// TIA Portal project "g" (V14)

(* hardware
DEVICE "S7-1200 station_1"  S7-1200 Station
   slot 0: "Rack_0"  S7-1200 Rack  Rack  V1.0
   slot 1: "PLC_1_test_mb_og_utv"  CPU 1217C DC/DC/DC  6ES7 217-1AG40-0XB0  V4.2
   slot 2: "DI 16x24VDC_1"  6ES7 221-1BH32-0XB0  V2.0
   slot 3: "CB 1241 (RS485)"  CB 1241 (RS485)  6ES7 241-1CH30-1XB0  V1.0
DEVICE "S7-1200 station_6"  S7-1200 Station
   slot 0: "Rack_0"  S7-1200 Rack  Rack  V1.0
   slot 1: "slib"  CPU 1211C DC/DC/DC  6ES7 211-1AE40-0XB0  V4.2
   slot 3: "CB 1241 (RS485)"  CB 1241 (RS485)  6ES7 241-1CH30-1XB0  V1.0
DEVICE "HMI"  TP900 Comfort
   slot 0: "TP900 Comfort"  TP900 Comfort  6AV2 124-0JC01-0AX0  14.0.1.0
   slot 1: "HMI_RT_2"  TP900 Comfort  6AV2 124-0JC01-0AX0  14.0.1.0
   slot 5: "HMI_2.IE_CP_1"  PROFINET Interface  14.0.1.0
      slot 1: "PROFINET Interface_1"  PROFINET Interface
         slot 1: "Port_1"  Port
         slot 2: "Port_2"  Port
   slot 7: "HMI_2.MPI/DP_CP_1"  MPI/DP Interface  14.0.1.0
DEVICE "S7-1200 station_2"  S7-1200 Station
   slot 0: "Rack_0"  S7-1200 Rack  Rack  V1.0
   slot 1: "PLC_1"  CPU 1211C DC/DC/DC  6ES7 211-1AE40-0XB0  V4.2
   slot 3: "CB 1241 (RS485)"  CB 1241 (RS485)  6ES7 241-1CH30-1XB0  V1.0
*)

// ===== PLC "PLC_1_test_mb_og_utv"  CPU 1217C DC/DC/DC =====

VAR_GLOBAL   // PLC tag table "Default tag table"
   "my_special_tag_name" AT %IW0 : Int;
   "tt" AT %I0.0 : Bool;
END_VAR

TYPE "mb_station_block_udt"
   STRUCT
      conf : Struct   // Configuration
         disable : Bool;   // Skip all queries
         read_only : Bool;   // Skip all write queries. (fc 5,6,15,16)
         max_comm_error : USInt := 2;   // Repeating erros before communication_error flag is set
         exec_x_quries : USInt := 1;   // Number of queries to be exec. at each loop.
      END_STRUCT;
      out : Struct   // Outputs
         error : Bool;   // All errors, including communication errors
         error_comm : Bool;   // only communication errors
         finnish : Bool;   // qid is handed over to next device.
      END_STRUCT;
      log : Struct   // Logging for development and debugging.
         connected_time : DTL;   // The time the device was connected to the bus
         disconnected_time : DTL;   // The time, if a device was disconnected to the bus
         done_cnt : UDInt;   // Successfully queries counter for this device
         error_comm_cnt : UDInt;   // Communication erros cnt.
         error_exception_cnt : UDInt;   // Failed queries counter for this device
         error_status : Word;   // Status code from mb_master or mb_client
         error_data_addr : UDInt;   // d_addr for last failed querie; handy for troubleshooting
      END_STRUCT;
      z : Struct   // Internal states.
         header_qid : UInt;   // qid value at device header
         comm_err_cnt : USInt;   // Repeating communication errors
         exec_cnt : USInt;   // Numb. of exec. q. this loop
         offset_qid : UInt := 1;   // Device query id.
         err_hold : Bool;   // Help var for .out.error
      END_STRUCT;
   END_STRUCT;
END_TYPE

// folder: mb_test

DATA_BLOCK "test_mb_t1_DB"   // DB1
{ S7_Optimized_Access := 'TRUE' }
VERSION : 0.1
// stored: InstanceOfName test_mb_1
"test_mb_1"
BEGIN
END_DATA_BLOCK

// folder: (top level)

FUNCTION_BLOCK "_read little"   // FB1, SCL
{ S7_Optimized_Access := 'TRUE' }
VERSION : 0.1
   VAR_INPUT
      mb_addr : USInt;
   END_VAR
   VAR_IN_OUT
      mb_query : "mb_query";
   END_VAR
   VAR
      sb : "mb_station_block_udt";
      data1 : Real;
      data2 : Real;
      data3 : Real;
      dommy : Bool;
      err : Int;
      pos : DInt;
   END_VAR
BEGIN

   #mb_query(mb_addr := 123,
             mode := #mb_query.c.read.holding_reg,
             data_addr := 12345,
             data_ptr := #dommy);

   IF #mb_query.Done THEN

       // #pos := "mb_pos"(mb_query := #mb_query, addr := 12345);
       #pos := UDINT_TO_DINT(12354 - #mb_query.data_addr) * 2;

       #err := READ_LITTLE(src_array := #mb_query.z.buffer,
                           dest_Variable => #data1,
                           pos := #pos);
       #err := READ_LITTLE(src_array := #mb_query.z.buffer,
                           dest_Variable => #data2,
                           pos := #pos);
       #err := READ_LITTLE(src_array := #mb_query.z.buffer,
                           dest_Variable => #data3,
                           pos := #pos);
   END_IF;
END_FUNCTION_BLOCK

FUNCTION_BLOCK "ABcounterEncoder"   // FB2, SCL
{ S7_Optimized_Access := 'TRUE' }
VERSION : 0.1
   VAR_INPUT
      pulsA : Bool;
      pulsB : Bool;
      reverce : Bool;
      factor : Real := 1.0;
   END_VAR
   VAR_OUTPUT
      pos : Real;
      uncertainPos : Bool;
   END_VAR
   VAR
      old : Struct
         pulsA : Bool;
         pulsB : Bool;
      END_STRUCT;
      cnt : DInt;
      firstScan : Bool := true;
   END_VAR
BEGIN
   // Position encoder based on two pulses which are 90 degree
   // phase shifted. 

   // TIP: Use a HSC (High speed conter) instead of this function
   // block. Using a hardware HSC will use less CPU resources.

   IF #firstScan THEN
       #uncertainPos := true;
   END_IF;

   IF #pulsA <> #old.pulsA OR #pulsB <> #old.pulsB THEN
       #cnt += SEL(G := #reverce XOR (
                    #pulsA <> NOT #old.pulsA
                    OR #pulsB <> NOT #old.pulsB),
                    IN0 := -1, IN1 := 1);
   END_IF;

   #pos := DINT_TO_REAL(#cnt) * #factor;
   #old.pulsA := #pulsA; 
   #old.pulsB := #pulsB; 
   #firstScan := false;
END_FUNCTION_BLOCK

FUNCTION_BLOCK "ABcounterCorrection"   // FB4, SCL
{ S7_Optimized_Access := 'TRUE' }
VERSION : 0.1
   VAR_INPUT
      switch : Bool;
      cnt : DInt;
   END_VAR
   VAR_OUTPUT
      deviation : DInt;
   END_VAR
   VAR_IN_OUT
      AB : "ABcounterEncoder";
   END_VAR
   VAR
      rtrig : R_TRIG;
   END_VAR
BEGIN
   #rtrig(CLK := #switch);

   // Log the max deviation
   IF NOT #AB.uncertainPos THEN
       #deviation := MAX(IN1 := #deviation, IN2 := ABS(#AB.cnt - #cnt));
   END_IF;

   IF #rtrig.Q THEN
       #AB.cnt := #cnt;
       #AB.uncertainPos := false;
   END_IF;
END_FUNCTION_BLOCK

FUNCTION "mb_get" : Void   // FC6, SCL
{ S7_Optimized_Access := 'TRUE' }
VERSION : 0.1
   VAR_INPUT
      addr : UDInt;
   END_VAR
   VAR_IN_OUT
      data_ptr : Variant;
      mb_query : "mb_query";
   END_VAR
   VAR_TEMP
      pos : DInt;
      err : Int;
   END_VAR
BEGIN
   IF #mb_query.z.run.qid_cnt = #mb_query.z.run.qid
       AND  #mb_query.Done
   THEN
       #pos := UDINT_TO_USINT(#addr - #mb_query.data_addr) * 2;
       #err := Deserialize(SRC_ARRAY := #mb_query.z.buffer,
                           DEST_VARIABLE => #data_ptr,
                           POS := #pos);
   END_IF;
END_FUNCTION

FUNCTION "mb_read_little_endian" : Void   // FC8, SCL
{ S7_Optimized_Access := 'TRUE' }
VERSION : 0.1
   VAR_INPUT
      addr : UDInt;
      n : USInt;
   END_VAR
   VAR_IN_OUT
      mb_query : "mb_query";
   END_VAR
   VAR_TEMP
      bo : Int;
      tmp : Byte;
      c : Int;
   END_VAR
BEGIN
   (* Read little endian:

      The function should be placed before a read query, and may be used 
      muliple times.

      "mb_read_little_endian"(addr := 100, n := 1, mb_query := #mb_query);
      "mb_read_little_endian"(addr := 200, n := 3, mb_query := #mb_query);

      #mb_query(mb_addr := ___MB_ADDR___,
                mode := #mb_query.c.read.holding_reg,
                data_addr := ___DATA_ADDR___,
                data_ptr := ___DATA___ );
   *) 

   IF #mb_query.z.run.qid_cnt + 1 = #mb_query.z.run.qid
       AND #mb_query.stat.done
       AND NOT #mb_query.z.run.insert
       AND NOT #mb_query.z.run.write // Read query
       AND #mb_query.conf.buffer_handler
   THEN
       #bo := UDINT_TO_INT(#addr - #mb_query.z.q.data_addr) * 2;

       FOR #c := #bo TO #bo + #n * 4 BY 4 DO
           #tmp := #mb_query.z.buffer[#bo + 0];
           #mb_query.z.buffer[#bo + 0] := #mb_query.z.buffer[#bo + 3];
           #mb_query.z.buffer[#bo + 3] := #tmp;

           #tmp := #mb_query.z.buffer[#bo + 1];
           #mb_query.z.buffer[#bo + 1] := #mb_query.z.buffer[#bo + 2];
           #mb_query.z.buffer[#bo + 2] := #tmp;
       END_FOR;
   END_IF;
END_FUNCTION

FUNCTION "mb_extra" : Bool   // FC9, SCL
{ S7_Optimized_Access := 'TRUE' }
VERSION : 0.1
   VAR_IN_OUT
      sb : "mb_station_block_udt";
      mb_query : "mb_query";
   END_VAR
BEGIN
   (* Example

   "mb_station_block_footer"(sb := #sb, mb_query := #mb_query);

   IF "mb_extra"(sb := #sb, mb_query := #mb_query) THEN
       #mb_query(mode := #mb_query.c.write.holding_reg,
                 data_addr := 12345,
                 data_ptr := ___CONFIG_PARAM___);
   END_IF;
   *)

   #mb_extra :=
   #mb_query.z.sb.sid = #mb_query.z.sb.sid_cnt
   AND NOT #sb.out.error_comm;
   // AND NOT #mb_query.stat.busy;
END_FUNCTION

ORGANIZATION_BLOCK "Main"   // OB1, SCL, ProgramCycle
TITLE = "Main Program Sweep (Cycle)"
{ S7_Optimized_Access := 'TRUE' }
VERSION : 0.1
   VAR_INPUT
      Initial_Call : Bool;   // Initial call of this OB
      Remanence : Bool;   // =True, if remanent data are available
   END_VAR
BEGIN
END_ORGANIZATION_BLOCK

// folder: mb_test

FUNCTION_BLOCK "test_mb_master"   // FB13, SCL
{ S7_Optimized_Access := 'TRUE' }
VERSION : 0.1
   VAR_INPUT
      REQ : Bool;
      MB_ADDR : UInt;
      MODE : USInt;
      DATA_ADDR : UDInt;
      DATA_LEN : UInt;
   END_VAR
   VAR_OUTPUT
      BUSY : Bool;
      ERROR : Bool;
      DONE : Bool;
      STATUS : Word;
   END_VAR
   VAR_IN_OUT
      DATA_PTR : "mb_internal_b";
   END_VAR
   VAR
      test : "test_mb_common";
   END_VAR
BEGIN
   #test(REQ := #REQ,
         MB_ADDR := #MB_ADDR,
         MODE := #MODE,
         DATA_ADDR := #DATA_ADDR,
         DATA_LEN := #DATA_LEN,
         BUSY => #BUSY,
         ERROR => #ERROR,
         DONE => #DONE,
         STATUS => #STATUS);
END_FUNCTION_BLOCK

FUNCTION_BLOCK "test_mb_common"   // FB14, SCL
{ S7_Optimized_Access := 'TRUE' }
VERSION : 0.1
   VAR_INPUT
      REQ : Bool;
      MB_ADDR : UInt;
      MODE : USInt;
      DATA_ADDR : UDInt;
      DATA_LEN : UInt;
   END_VAR
   VAR_OUTPUT
      BUSY : Bool;
      ERROR : Bool;
      DONE : Bool;
      STATUS : Word;
   END_VAR
   VAR
      fakeBus : Struct
         q : Struct
            mb_addr : UInt;
            mode : USInt;
            data_addr : UDInt;
            data_len : UInt;
         END_STRUCT;
         res : Struct
            done : Bool;
            error : Bool;
         END_STRUCT;
      END_STRUCT;
      state : Int;
      reset : Bool;
      cnt : Int;
   END_VAR
BEGIN
   // Fake query testing block

   CASE #state OF
       0:  // Wait for req.
           IF #REQ THEN
               #BUSY := true;
               #state += 1;
           END_IF;
           #cnt := 0; // Init cnt.

       1:  // Simulate some waite time
           #cnt += 1;
           #state += BOOL_TO_INT(#cnt > 5);

       2:  // Insert q-param to fake bus.
           #fakeBus.q.mb_addr := #MB_ADDR;
           #fakeBus.q.mode := #MODE;
           #fakeBus.q.data_addr := #DATA_ADDR;
           #fakeBus.q.data_len := #DATA_LEN;
           #cnt += 1; // The test device will insert resualt until next scan.

       3:  // Done or Eroor
           #fakeBus.q.mb_addr := 0;
           #fakeBus.q.mode := 0;
           #fakeBus.q.data_addr := 0;
           #fakeBus.q.data_len := 0;

           #DONE := #fakeBus.res.done;
           #ERROR := #fakeBus.res.error;
           IF NOT #DONE AND NOT #ERROR THEN
               #ERROR := true;
               #STATUS := 16#80C8;
           END_IF;
           #BUSY := false;
           #state := 0;
   END_CASE;

   IF #reset THEN
       #state := 0;
       #ERROR := false;
       #DONE := false;
       #BUSY := false;
   END_IF;

   #fakeBus.res.done := false;
   #fakeBus.res.error := false;
END_FUNCTION_BLOCK

FUNCTION_BLOCK "test_mb_client"   // FB15, SCL
{ S7_Optimized_Access := 'TRUE' }
VERSION : 0.1
   VAR_INPUT
      REQ : Bool;
      DISCONNECT : Bool;
      MB_MODE : USInt;
      DATA_ADDR : UDInt;
      DATA_LEN : UInt;
   END_VAR
   VAR_OUTPUT
      DONE : Bool;
      BUSY : Bool;
      ERROR : Bool;
      STATUS : Word;
   END_VAR
   VAR_IN_OUT
      MB_DATA_PTR : Variant;
      CONNECT : Variant;
   END_VAR
   VAR
      MB_Unit_ID : USInt;
      Connected : Bool;
      _ : Bool;
      test : "test_mb_common";
      cnt : UInt;
   END_VAR
BEGIN
   IF #DISCONNECT THEN
       #cnt := 0;
       #test.reset := true;
       #Connected := false;
   ELSE
       IF #cnt < 10 THEN
           #cnt += 1;
           #BUSY := true;
       ELSE
           #Connected := true;
           #test.reset := false;

       END_IF;
   END_IF;

   #test(REQ := #REQ,
         MB_ADDR := #MB_Unit_ID,
         MODE := #MB_MODE,
         DATA_ADDR := #DATA_ADDR,
         DATA_LEN := #DATA_LEN,
         BUSY => #BUSY,
         ERROR => #ERROR,
         DONE => #DONE,
         STATUS => #STATUS);
END_FUNCTION_BLOCK

FUNCTION_BLOCK "test_mb_1"   // FB16, SCL
{ S7_Optimized_Access := 'TRUE' }
VERSION : 0.1
   VAR_INPUT
      start : Bool;
   END_VAR
   VAR_OUTPUT
      DONE : Bool;
      ERROR : Bool;
   END_VAR
   VAR
      state : Int;
      old_state : Int;
      cnt : UInt;
      mx : UInt;
      mb_query : "mb_query";
      mb_master_1200_ctrl : "mb_master_1200_ctrl";
      mb_master_1500_ctrl : "mb_master_1200_ctrl";
      mb_client_ctrl : "mb_client_ctrl";
      mb_test_sb : Array[1..5] of "test_mb_sb1";
      mb_test_sb_fake : Array[1..5] of "test_mb_sb1_fake_device";
   END_VAR
   VAR_TEMP
      c : Int;
      dommy : Word;
   END_VAR
BEGIN
   CASE #state OF
       0:  // Wait for start signal.
           #state += BOOL_TO_INT(#start);
           #DONE := false;
           #ERROR := false;

       1:  // mb_master-1200
           #mb_test_sb[1].write1.real_1 := 0;
           #mb_test_sb[1].write1.real_2 := 0;
           #mb_test_sb[4].write1.real_1 := 0;
           #mb_test_sb[4].write1.real_2 := 0;
           #state += 1;
       2:  
           #mb_master_1200_ctrl(hardware_id := 1,
                                baud := 9600,
                                timeout := T#0s, // Auto
                                mb_query := #mb_query);

           #mb_test_sb[1].write1.real_1 := 12.34;
           #mb_test_sb[1].write1.real_2 := 56.78;
           #mb_test_sb[1]<?Sub?>(MB_ADDR := 1, mb_query := #mb_query);
           #mb_test_sb[2]<?Sub?>(MB_ADDR := 1, mb_query := #mb_query);
           #mb_test_sb[3]<?Sub?>(MB_ADDR := 1, mb_query := #mb_query);

           // Create some noice ...
           FOR #c := 0 TO UINT_TO_INT( #cnt ) MOD 7 DO
               #mb_query(mb_addr := 200, data_ptr := #dommy);
           END_FOR;

           #mb_test_sb[4].write1.real_1 := 90.12;
           #mb_test_sb[4].write1.real_2 := 34.56;
           #mb_test_sb[4]<?Sub?>(MB_ADDR := 1, mb_query := #mb_query);
           #mb_test_sb[5]<?Sub?>(MB_ADDR := 1, mb_query := #mb_query);

           FOR #c := 1 TO 5 DO
               #mb_test_sb_fake[#c]<?Sub?>(MB_ADDR := INT_TO_USINT(#c),
                                    mb_query := #mb_query,
                                    mb_test := #mb_master_1200_ctrl.master.TEST,
                                    mb_buffer := #mb_master_1200_ctrl.buffer.buffer);
           END_FOR;

           #state += BOOL_TO_INT(#cnt > 10000
                                 AND #mb_test_sb[1].read1.real_1 <> 12.34
                                 AND #mb_test_sb[1].read1.real_2 <> 56.78
                                 AND #mb_test_sb[4].read1.real_1 <> 90.12
                                 AND #mb_test_sb[4].read1.real_2 <> 34.56 );

           IF #mb_test_sb[1].read1.real_1 <> 12.34 AND #mb_test_sb[1].read1.real_1 <> 0
               OR #mb_test_sb[1].read1.real_2 <> 56.78 AND #mb_test_sb[1].read1.real_2 <> 0

               OR #mb_test_sb[4].read1.real_1 <> 90.12 AND #mb_test_sb[4].read1.real_1 <> 0
               OR #mb_test_sb[4].read1.real_2 <> 34.56 AND #mb_test_sb[4].read1.real_2 <> 0
           THEN
               #state := -1; // Error
           END_IF;

       3:  // 1500
           #mb_test_sb[3].read1.real_1 := 0;
           #state += 1;
       4:
           #mb_master_1500_ctrl(hardware_id := 1,
                                baud := 9600,
                                timeout := T#300ms,
                                mb_query := #mb_query);

           #mb_test_sb[3].write1.real_1 := 98.76;

           FOR #c := 1 TO 5 DO
               #mb_test_sb[#c]<?Sub?>(MB_ADDR := INT_TO_USINT(#c),
                               mb_query := #mb_query);
           END_FOR;

           #mb_test_sb_fake[2]<?Sub?>(MB_ADDR := INT_TO_USINT(2),
                               mb_query := #mb_query,
                               mb_test := #mb_master_1500_ctrl.master.TEST,
                               mb_buffer := #mb_master_1500_ctrl.buffer.buffer);

           #state += BOOL_TO_INT(#cnt > 10000 AND #mb_test_sb[3].read1.real_1 <> 98.76 );

           IF #mb_test_sb[3].read1.real_1 <> 98.76 AND #mb_test_sb[3].read1.real_1 <> 0 THEN
               #state := -2; // Error
               #state += 1;
           END_IF;

       5:  // Client
           #mb_test_sb[2].read1.real_1 := 0;
       6:
           #mb_client_ctrl(mb_query := #mb_query);

           #mb_test_sb[2].write1.real_1 := 0.000076;

           FOR #c := 1 TO 5 DO
               #mb_test_sb[#c]<?Sub?>(MB_ADDR := INT_TO_USINT(#c), mb_query := #mb_query);
           END_FOR;

           #mb_test_sb_fake[2]<?Sub?>(MB_ADDR := INT_TO_USINT(2),
                               mb_query := #mb_query,
                               mb_test := #mb_master_1200_ctrl.master.TEST,
                               mb_buffer := #mb_master_1200_ctrl.buffer.buffer);

           #state += BOOL_TO_INT(#cnt > 10000
                                 AND #mb_test_sb[2].read1.real_1 <> 0.000076);

           IF #mb_test_sb[2].read1.real_1 <> 0.000076 AND #mb_test_sb[2].read1.real_1 <> 0 THEN
               #state := -2; // Error
           END_IF;

       7:
           #DONE := true;
   END_CASE;

   #cnt += 1;
   IF #old_state <> #state THEN
       #cnt := 0;
   END_IF;
   #old_state := #state;

   #ERROR := #state < 0;
END_FUNCTION_BLOCK

FUNCTION_BLOCK "test_mb_comm_load"   // FB17, SCL
{ S7_Optimized_Access := 'TRUE' }
VERSION : 0.1
   VAR_INPUT
      REQ : Bool;
      PORT : Port;
      BAUD : UInt;
      PARITY : UInt;
      RESP_TO : UInt;
   END_VAR
   VAR_OUTPUT
      DONE : Bool;
      ERROR : Bool;
   END_VAR
   VAR_IN_OUT
      MB_DB : Variant;
   END_VAR
   VAR
      MB_COMM_LOAD_Instance : MB_COMM_LOAD;
      "1500" : Bool;
   END_VAR
BEGIN

   IF #"1500" THEN
       #DONE := false;
   END_IF;

   IF #REQ  
       AND #PORT <> 0 AND #BAUD <> 0 AND #PARITY <> 0 AND #RESP_TO <> 0
   THEN
       #DONE := true;
   END_IF;

   #ERROR := NOT #DONE;
END_FUNCTION_BLOCK

FUNCTION_BLOCK "test_mb_sb1_fake_device"   // FB18, SCL
{ S7_Optimized_Access := 'TRUE' }
VERSION : 0.1
   VAR_INPUT
      MB_ADDR : UInt;
   END_VAR
   VAR_IN_OUT
      mb_query : "mb_query";
      mb_test : "test_mb_common";
      mb_buffer : Array[0..250] of Byte;
   END_VAR
   VAR
      fakeBus : Struct
         q : Struct
            mb_addr : UInt;
            mode : USInt;
            data_addr : UDInt;
            data_len : UInt;
         END_STRUCT;
         res : Struct
            done : Bool;
            error : Bool;
         END_STRUCT;
      END_STRUCT;
      read1 : Struct
         real_1 : Real;
         real_2 : Real;
         udint_1 : UDInt;
      END_STRUCT;
      read2 : Struct
         x00 : Bool;
         x01 : Bool;
         x02 : Bool;
         x03 : Bool;
         x04 : Bool;
         x05 : Bool;
         x06 : Bool;
         x07 : Bool;
         x08 : Bool;
         x09 : Bool;
         x10 : Bool;
         x11 : Bool;
         x12 : Bool;
         x13 : Bool;
         x14 : Bool;
         x15 : Bool;
      END_STRUCT;
      write1 : Struct
         real_2 : Real;
         udint_1 : UDInt;
         real_1 : Real;
      END_STRUCT;
      sb : "mb_station_block_udt";
   END_VAR
   VAR_TEMP
      pos : DInt;
      "e" : Int;
   END_VAR
BEGIN
   // Simulating a device 

   IF #mb_test.fakeBus.q.mb_addr = #MB_ADDR 
       AND #mb_test.fakeBus.q.data_len > 1
   THEN
       // Read 1
       IF #mb_test.fakeBus.q.mode = #mb_query.c.read.holding_reg
           AND #mb_test.fakeBus.q.data_addr = 123
       THEN
           #"e" := Serialize(SRC_VARIABLE := #read1, DEST_ARRAY => #mb_buffer, POS := #pos);
           #mb_test.fakeBus.res.done := #"e" = 0 AND #pos / 2 = #mb_test.fakeBus.q.data_len;
       END_IF;

       // Read 2
       IF #mb_test.fakeBus.q.mode = #mb_query.c.read.holding_reg
           AND #mb_test.fakeBus.q.data_addr = 456
       THEN
           #"e" := Serialize(SRC_VARIABLE := #read2, DEST_ARRAY => #mb_buffer, POS := #pos);
           #mb_test.fakeBus.res.done := #"e" = 0 AND #pos / 2 = #mb_test.fakeBus.q.data_len;
       END_IF;

       // Write 1
       IF #mb_test.fakeBus.q.mode = #mb_query.c.write.holding_reg
           AND #mb_test.fakeBus.q.data_addr = 789
       THEN
           #"e" := Deserialize(SRC_ARRAY := #mb_buffer, DEST_VARIABLE => #write1, POS := #pos);
           #mb_test.fakeBus.res.done := #"e" = 0 AND #pos / 2 = #mb_test.fakeBus.q.data_len;
       END_IF;
   END_IF;

   #mb_test.fakeBus.res.error := NOT #mb_test.fakeBus.res.done;

   #read1.real_1 := #write1.real_1;
   #read1.real_2 := #write1.real_2;
   #read1.udint_1 := #write1.udint_1;
END_FUNCTION_BLOCK

FUNCTION_BLOCK "test_mb_sb1"   // FB19, SCL
{ S7_Optimized_Access := 'TRUE' }
VERSION : 0.1
   VAR_INPUT
      MB_ADDR : UInt;
   END_VAR
   VAR_IN_OUT
      mb_query : "mb_query";
   END_VAR
   VAR
      fakeBus : Struct
         q : Struct
            mb_addr : UInt;
            mode : USInt;
            data_addr : UDInt;
            data_len : UInt;
         END_STRUCT;
         res : Struct
            done : Bool;
            error : Bool;
         END_STRUCT;
      END_STRUCT;
      read1 : Struct
         real_1 : Real;
         real_2 : Real;
         udint_1 : UDInt;
      END_STRUCT;
      read2 : Struct
         x00 : Bool;
         x01 : Bool;
         x02 : Bool;
         x03 : Bool;
         x04 : Bool;
         x05 : Bool;
         x06 : Bool;
         x07 : Bool;
         x08 : Bool;
         x09 : Bool;
         x10 : Bool;
         x11 : Bool;
         x12 : Bool;
         x13 : Bool;
         x14 : Bool;
         x15 : Bool;
      END_STRUCT;
      write1 : Struct
         real_2 : Real;
         udint_1 : UDInt;
         real_1 : Real;
      END_STRUCT;
      sb : "mb_station_block_udt";
      q1_done_cnt : UDInt;
      q2_done_cnt : UDInt;
      q3_done_cnt : UDInt;
   END_VAR
BEGIN
   // Testing device

   "mb_station_block_header"(sb := #sb, mb_query := #mb_query);
   #mb_query.mb_addr := #MB_ADDR;

   #mb_query(mode := #mb_query.c.read.holding_reg,
             data_addr := 123,
             data_ptr := #read1);
   #q1_done_cnt += BOOL_TO_UDINT(#mb_query.Done);

   #mb_query(mode := #mb_query.c.read.holding_reg,
             data_addr := 456,
             data_ptr := #read2);
   #q2_done_cnt += BOOL_TO_UDINT(#mb_query.Done);

   #mb_query(mode := #mb_query.c.write.holding_reg,
             data_addr := 789,
             data_ptr := #write1);
   #q3_done_cnt += BOOL_TO_UDINT(#mb_query.Done);

   "mb_station_block_footer"(sb := #sb, mb_query := #mb_query);
END_FUNCTION_BLOCK

FUNCTION_BLOCK "test_mb_sb2"   // FB20, SCL
{ S7_Optimized_Access := 'TRUE' }
VERSION : 0.1
   VAR_INPUT
      MB_ADDR : UInt;
   END_VAR
   VAR_IN_OUT
      mb_query : "mb_query";
   END_VAR
   VAR
      fakeBus : Struct
         q : Struct
            mb_addr : UInt;
            mode : USInt;
            data_addr : UDInt;
            data_len : UInt;
         END_STRUCT;
         res : Struct
            done : Bool;
            error : Bool;
         END_STRUCT;
      END_STRUCT;
      read1 : Struct
         real_1 : Real;
         real_2 : Real;
         udint_1 : UDInt;
      END_STRUCT;
      read2 : Struct
         x00 : Bool;
         x01 : Bool;
         x02 : Bool;
         x03 : Bool;
         x04 : Bool;
         x05 : Bool;
         x06 : Bool;
         x07 : Bool;
         x08 : Bool;
         x09 : Bool;
         x10 : Bool;
         x11 : Bool;
         x12 : Bool;
         x13 : Bool;
         x14 : Bool;
         x15 : Bool;
      END_STRUCT;
      write1 : Struct
         real_2 : Real;
         udint_1 : UDInt;
         real_1 : Real;
      END_STRUCT;
      sb : "mb_station_block_udt";
      q1_done_cnt : UDInt;
      q2_done_cnt : UDInt;
      q3_done_cnt : UDInt;
   END_VAR
BEGIN
   // Testing device

   "mb_station_block_header"(sb := #sb, mb_query := #mb_query);
   #mb_query.mb_addr := #MB_ADDR;

   #mb_query(mode := #mb_query.c.read.holding_reg,
             data_addr := 123,
             data_ptr := #read1);
   #q1_done_cnt += BOOL_TO_UDINT(#mb_query.Done);

   #mb_query(mode := #mb_query.c.read.holding_reg,
             data_addr := 456,
             data_ptr := #read2);
   #q2_done_cnt += BOOL_TO_UDINT(#mb_query.Done);

   #mb_query(mode := #mb_query.c.write.holding_reg,
             data_addr := 789,
             data_ptr := #write1);
   #q3_done_cnt += BOOL_TO_UDINT(#mb_query.Done);

   "mb_station_block_footer"(sb := #sb, mb_query := #mb_query);
END_FUNCTION_BLOCK

FUNCTION_BLOCK "test_mb_sb2_fake_device"   // FB21, SCL
{ S7_Optimized_Access := 'TRUE' }
VERSION : 0.1
   VAR_INPUT
      MB_ADDR : UInt;
   END_VAR
   VAR_IN_OUT
      mb_query : "mb_query";
      mb_test : "test_mb_common";
      mb_buffer : Array[0..250] of Byte;
   END_VAR
   VAR
      fakeBus : Struct
         q : Struct
            mb_addr : UInt;
            mode : USInt;
            data_addr : UDInt;
            data_len : UInt;
         END_STRUCT;
         res : Struct
            done : Bool;
            error : Bool;
         END_STRUCT;
      END_STRUCT;
      read1 : Struct
         real_1 : Real;
         real_2 : Real;
         udint_1 : UDInt;
      END_STRUCT;
      read2 : Struct
         x00 : Bool;
         x01 : Bool;
         x02 : Bool;
         x03 : Bool;
         x04 : Bool;
         x05 : Bool;
         x06 : Bool;
         x07 : Bool;
         x08 : Bool;
         x09 : Bool;
         x10 : Bool;
         x11 : Bool;
         x12 : Bool;
         x13 : Bool;
         x14 : Bool;
         x15 : Bool;
      END_STRUCT;
      write1 : Struct
         real_2 : Real;
         udint_1 : UDInt;
         real_1 : Real;
      END_STRUCT;
      sb : "mb_station_block_udt";
   END_VAR
   VAR_TEMP
      pos : DInt;
      "e" : Int;
   END_VAR
BEGIN
   // Simulating a device 

   IF #mb_test.fakeBus.q.mb_addr = #MB_ADDR 
       AND #mb_test.fakeBus.q.data_len > 1
   THEN

       IF #mb_test.fakeBus.q.mode = #mb_query.c.read.input_reg
           AND #mb_test.fakeBus.q.data_addr = 123
       THEN
           #mb_test.fakeBus.res.done := false;
           #mb_test.STATUS := 16#8380; // CRC error 
       END_IF;

       IF #mb_test.fakeBus.q.mode = #mb_query.c.read.input_reg
           AND #mb_test.fakeBus.q.data_addr = 456
       THEN
           #mb_test.fakeBus.res.done := false;
           #mb_test.STATUS := 16#8384; // Data value error
       END_IF;

   END_IF;

   #mb_test.fakeBus.res.error := NOT #mb_test.fakeBus.res.done;

   #read1.real_1 := #write1.real_1;
   #read1.real_2 := #write1.real_2;
   #read1.udint_1 := #write1.udint_1;

   (* 

   Communications and configuration error messages of the instruction
   0000  No error
   80C8  Slave timeout. Check the baud rate, parity and the connectors on the slave.
   80D1  The receiver issued a flow control request to suspend an active transmission 
         and never re-enabled the transmission within the wait time.
   This  error is also generated during hardware flow control if the recipient does 
         not detect CTS within the wait time.
   80D2  The send request was aborted because no DSR signal is received from the DCE.
   80E0  The message was terminated because the receive buffer is full.
   80E1  The message was terminated as a result of a parity error.
   80E2  The message was terminated as a result of a framing error.
   80E3  The message was terminated as a result of an overrun error.
   80E4  The message was terminated as a result of the specified length exceeding the 
         total buffer size.
   8180  Invalid value for the port ID.
   8186  Invalid Modbus station address
   8188  The MODE parameter has an invalid value for a broadcast call.
   8189  Invalid data address value.
   818A  Invalid data length value.
   818B  Invalid pointer to the local data source/destination: Size not correct
   818C  The DATA_PTR parameter has an invalid pointer. Use a pointer to a bit memory 
         area or a DB with the "Standard - compatible with S7-300/400" access type.
   8200  Port is busy processing a send request


   Error messages of the Modbus protocol
   8380       CRC error 
   8381   01  Function code not supported
   8382   03  Data length error
   8383   02  Error in the data address or address outside the valid range of DATA_PTR
   8384  >03  Data value error
   8385   03  Data diagnostic code value not supported (function code 08)
   8386       Function code of the response does not match the function code of the query.
   8387       Response from wrong slave
   8388       The response of the slave to a write call is not correct. The data sent by 
              the slave does not match the query from the master.

   *)
END_FUNCTION_BLOCK

ORGANIZATION_BLOCK "test_mb_main_OB"   // OB123, SCL, ProgramCycle
TITLE = "Main Program Sweep (Cycle)"
{ S7_Optimized_Access := 'TRUE' }
VERSION : 0.1
   VAR_INPUT
      Initial_Call : Bool;   // Initial call of this OB
      Remanence : Bool;   // =True, if remanent data are available
   END_VAR
BEGIN
   "test_mb_t1_DB"();
END_ORGANIZATION_BLOCK

// ===== PLC "slib"  CPU 1211C DC/DC/DC =====

VAR_GLOBAL CONSTANT   // PLC tag table "Default tag table"
   "Handshakes.iSize" : Int := 10;
END_VAR

// folder: Library/Modbus/Core/sb

TYPE "mb_station_block_udt"
   STRUCT
      conf : Struct   // Configuration
         skip_code : Bool;
         disable : Bool;   // Skip all queries
         read_only : Bool;   // Skip all write queries. (fc 5,6,15,16)
         max_comm_error : USInt := 2;   // Repeating erros before communication_error flag is set
         exec_x_quries : USInt := 1;   // Number of queries to be exec. at each loop.
      END_STRUCT;
      out : Struct   // Outputs
         error : Bool;   // All errors, including communication errors
         error_comm : Bool;   // only communication errors
         finnish : Bool;   // qid is handed over to next device.
      END_STRUCT;
      log : Struct   // Logging for development and debugging.
         connected_time : DTL;   // The time the device was connected to the bus
         disconnected_time : DTL;   // The time, if a device was disconnected to the bus
         done_cnt : UDInt;   // Successfully queries counter for this device
         error_comm_cnt : UDInt;   // Communication erros cnt.
         error_exception_cnt : UDInt;   // Failed queries counter for this device
         error_status : Word;   // Status code from mb_master or mb_client
         error_data_addr : UDInt;   // d_addr for last failed querie; handy for troubleshooting
      END_STRUCT;
      z : Struct   // Internal states.
         header_qid : UInt;   // qid value at device header
         comm_err_cnt : USInt;   // Repeating communication errors
         exec_cnt : USInt;   // Numb. of exec. q. this loop
         offset_qid : UInt := 1;   // Device query id.
         err_hold : Bool;   // Help var for .out.error
      END_STRUCT;
   END_STRUCT;
END_TYPE

// ===== PLC "PLC_1"  CPU 1211C DC/DC/DC =====

// folder: Library/Modbus/Core/sb

TYPE "mb_station_block_udt"
   STRUCT
      conf : Struct   // Configuration
         skip_code : Bool;
         disable : Bool;   // Skip all queries
         read_only : Bool;   // Skip all write queries. (fc 5,6,15,16)
         max_comm_error : USInt := 2;   // Repeating erros before communication_error flag is set
         exec_x_quries : USInt := 1;   // Number of queries to be exec. at each loop.
      END_STRUCT;
      out : Struct   // Outputs
         error : Bool;   // All errors, including communication errors
         error_comm : Bool;   // only communication errors
         finnish : Bool;   // qid is handed over to next device.
      END_STRUCT;
      log : Struct   // Logging for development and debugging.
         connected_time : DTL;   // The time the device was connected to the bus
         disconnected_time : DTL;   // The time, if a device was disconnected to the bus
         done_cnt : UDInt;   // Successfully queries counter for this device
         error_comm_cnt : UDInt;   // Communication erros cnt.
         error_exception_cnt : UDInt;   // Failed queries counter for this device
         error_status : Word;   // Status code from mb_master or mb_client
         error_data_addr : UDInt;   // d_addr for last failed querie; handy for troubleshooting
      END_STRUCT;
      z : Struct   // Internal states.
         header_qid : UInt;   // qid value at device header
         comm_err_cnt : USInt;   // Repeating communication errors
         exec_cnt : USInt;   // Numb. of exec. q. this loop
         offset_qid : UInt := 1;   // Device query id.
         err_hold : Bool;   // Help var for .out.error
      END_STRUCT;
   END_STRUCT;
END_TYPE

// folder: Library/Modbus/Station blocks/Mettler

TYPE "mettlerToledoInd560Udt"
   STRUCT
      readMsgSlot : Array[1..4] of Struct
         cmdRespons : Struct
            FP_1 : Bool;
            FP_2 : Bool;
            FP_3 : Bool;
            FP_4 : Bool;
            FP_5 : Bool;
            data_integrity : Bool;
            cmdAck1 : Bool;
            cmdAck2 : Bool;
         END_STRUCT;
         reserved : Byte;   // volt
         data : Real;
         scale_status : Struct
            x08_Enter_Key : Bool;
            x09_Input_1 : Bool;
            x10_Input_2 : Bool;
            x11_Input_3 : Bool;
            x12_Motion : Bool;
            x13_Net_Mode : Bool;
            x14_Data_Integrity_2 : Bool;
            x15_Data_OK : Bool;
            x00_Target_1 : Bool;
            x01_Comparator_1 : Bool;
            x02_Targe_2 : Bool;
            x03_Comparator_2 : Bool;
            x04_Target_3 : Bool;
            x05_Alway_true : Bool;
            x06_TE_bit_1 : Bool;
            x07_TE_bit_2 : Bool;
         END_STRUCT;
      END_STRUCT;
      writeMsgSlot : Array[1..4] of Struct
         cmd : UInt;
         data : Real;
      END_STRUCT;
      run : Struct   // Data calculated from readMsgSlot
         PF : Array[1..4] of USInt;   // Floating point input indication
         cmdAck : Array[1..4] of USInt;
      END_STRUCT;
      occupiedMsgSlots : Array[1..4] of Bool;
      queryDone : Struct
         read : Bool;
         write : Bool;
      END_STRUCT;
   END_STRUCT;
END_TYPE

// folder: (top level)

FUNCTION_BLOCK "modbus_test_rtu_1200"   // FB3, SCL
{ S7_Optimized_Access := 'TRUE' }
VERSION : 0.1
   VAR
      mb_query : "mb_query";
      mb_master_1200_ctrl : "mb_master_1200_ctrl";
      delay_between_queries : "mb_delay_between_queries";
      delay : "mb_delay";
      __ : Bool;
      temperature_1 : "Jdrk_RS_WS_N01_1";
      temperature_2 : "Jdrk_RS_WS_N01_1";
      temperature_3 : "Jdrk_RS_WS_N01_1";
      sb_temp_no_answer_1 : "sb_temp_no_answer_1";
      sb_temp_no_answer_2 : "sb_temp_no_answer_1";
      sb_temp_no_answer_3 : "sb_temp_no_answer_1";
      sb_temp_error_1 : "sb_temp_error_1";
      sb_temp_error_2 : "sb_temp_error_1";
      sb_temp_error_3 : "sb_temp_error_1";
      _ : Bool;
      bool_arrary : Array[0..15] of Bool;
      sb : "mb_station_block_udt";
   END_VAR
BEGIN
   #mb_master_1200_ctrl.conf.parity := 0;
   #mb_master_1200_ctrl(hardware_id := 269, // "Local~CB_1241_(RS485)",
                        baud := 9600,
                        mb_query := #mb_query);

   #delay_between_queries(mb_query :=#mb_query);

   #temperature_1(mb_query := #mb_query);
   #temperature_2(mb_query := #mb_query);
   #temperature_3(mb_query := #mb_query);

   #delay(mb_query := #mb_query);

   #sb_temp_no_answer_1(mb_query := #mb_query);
   #sb_temp_no_answer_2(mb_query := #mb_query);
   #sb_temp_no_answer_3(mb_query := #mb_query);

   #sb_temp_error_1(mb_query := #mb_query);
   #sb_temp_error_2(mb_query := #mb_query);
   #sb_temp_error_3(mb_query := #mb_query);

   "mb_station_block_header"(sb := #sb, mb_query := #mb_query);
   #mb_query.mb_addr := 1;
   #mb_query.mode := #mb_query.c.read.input_reg;
   #mb_query.data_addr := 1;
   "mb_query_bits"(data_ptr := #bool_arrary, mb_query := #mb_query);
   "mb_station_block_footer"(sb := #sb, mb_query := #mb_query);
END_FUNCTION_BLOCK

FUNCTION_BLOCK "sb_temp_no_answer_1"   // FB4, SCL
{ S7_Optimized_Access := 'TRUE' }
VERSION : 0.1
   VAR_OUTPUT
      Temperature : Real;
   END_VAR
   VAR_IN_OUT
      mb_query : "mb_query";
   END_VAR
   VAR
      sb : "mb_station_block_udt";
   END_VAR
   VAR RETAIN
      offset : Real;
   END_VAR
   VAR_TEMP
      tmp : Int;
   END_VAR
BEGIN
   // JDRK - RS-WS-N01-8 - Temperature and Humidity sensor

   "mb_station_block_header"(sb := #sb, mb_query := #mb_query);

   #mb_query(mb_addr := 200,
             mode := #mb_query.c.read.input_reg,
             data_addr := 1,
             data_ptr := #tmp);

   IF #mb_query.Done THEN
       #Temperature := INT_TO_REAL(#tmp) / 10 + #offset;
   END_IF;

   "mb_station_block_footer"(sb := #sb, mb_query := #mb_query);
END_FUNCTION_BLOCK

FUNCTION_BLOCK "Jdrk_RS_WS_N01_1"   // FB31, SCL
{ S7_Optimized_Access := 'TRUE' }
VERSION : 0.1
   VAR_OUTPUT
      Temperature : Real;
   END_VAR
   VAR_IN_OUT
      mb_query : "mb_query";
   END_VAR
   VAR
      sb : "mb_station_block_udt";
   END_VAR
   VAR RETAIN
      offset : Real;
   END_VAR
   VAR_TEMP
      tmp : Int;
   END_VAR
BEGIN
   // JDRK - RS-WS-N01-8 - Temperature and Humidity sensor

   "mb_station_block_header"(sb := #sb, mb_query := #mb_query);

   #mb_query(mb_addr := 1,
             mode := #mb_query.c.read.input_reg,
             data_addr := 1,
             data_ptr := #tmp);

   IF #mb_query.Done THEN
       #Temperature := INT_TO_REAL(#tmp) / 10 + #offset;
   END_IF;

   "mb_station_block_footer"(sb := #sb, mb_query := #mb_query);
END_FUNCTION_BLOCK

FUNCTION_BLOCK "sb_temp_error_1"   // FB33, SCL
{ S7_Optimized_Access := 'TRUE' }
VERSION : 0.1
   VAR_OUTPUT
      Temperature : Real;
   END_VAR
   VAR_IN_OUT
      mb_query : "mb_query";
   END_VAR
   VAR
      sb : "mb_station_block_udt";
   END_VAR
   VAR RETAIN
      tt : Array[0..100] of Int;
   END_VAR
   VAR_TEMP
      tmp : Int;
   END_VAR
BEGIN
   // JDRK - RS-WS-N01-8 - Temperature and Humidity sensor

   "mb_station_block_header"(sb := #sb, mb_query := #mb_query);

   #mb_query(mb_addr := 1,
             mode := #mb_query.c.read.input_reg,
             data_addr := 1,
             data_ptr := #tmp);

   IF #mb_query.Done THEN
       #Temperature := INT_TO_REAL(#tmp) / 10;
   END_IF;

   // Query producing a error.
   #mb_query(mb_addr := 1,
             mode := #mb_query.c.read.input_reg,
             data_addr := 1,
             data_ptr := #tt);

   "mb_station_block_footer"(sb := #sb, mb_query := #mb_query);
END_FUNCTION_BLOCK

ORGANIZATION_BLOCK "Main"   // OB1, SCL, ProgramCycle
TITLE = "Main Program Sweep (Cycle)"
{ S7_Optimized_Access := 'TRUE' }
VERSION : 0.1
   VAR_INPUT
      Initial_Call : Bool;   // Initial call of this OB
      Remanence : Bool;   // =True, if remanent data are available
   END_VAR
BEGIN
END_ORGANIZATION_BLOCK

// folder: Library/Modbus/Core

FUNCTION_BLOCK "mb_query"   // FB1, SCL
{ S7_Optimized_Access := 'TRUE' }
VERSION : 0.1
   VAR_INPUT
      mb_addr : UInt;   // Device addr. (0 to 247)
      mode : USInt;   // Function code: 1,2,3,4,5,6,15,16. (siemens mode shifted to 200 - 202)
      data_addr : UDInt;   // Data addr. (raw telegram value, 0-65535)
      data_len : UInt;   // Data len. 0=>Auto detect
   END_VAR
   VAR_OUTPUT
      Done : Bool;   // Successful query
      Error : Bool;   // Failed query
   END_VAR
   VAR_IN_OUT
      data_ptr : Variant;   // Bytes and bools has to add up to whole word(s)
   END_VAR
   VAR
      c : Struct   // Constants
         read : Struct   // Read: 1, 2, 3, 4
            discrete_output : USInt := 1;   // 1 (coils)
            discrete_input : USInt := 2;   // 2
            holding_reg : USInt := 3;   // 3
            input_reg : USInt := 4;   // 4
         END_STRUCT;
         write : Struct   // Write: 5, 6, 15, 16
            single_discrete_output : USInt := 5;   // 5 (coil) (when len. is eq. to 1)
            single_holding_reg : USInt := 6;   // 6 (when len. is eq. to 1)
            discrete_output : USInt := 15;   // 15 (coils)
            holding_reg : USInt := 16;   // 16
         END_STRUCT;
         mode : Struct   // Modicon convention addressing. (Eg: hold.reg. start at 40001)
            read : USInt := 200;   // Mode 0 (fc: 1, 2, 3, 4)
            write_single : USInt := 201;   // Mode 1 (fc: 5, 6) (when len. is eq. to 1)
            write : USInt := 202;   // Mode 2 (fc: 15, 16)
         END_STRUCT;
         auto_len : USInt := 0;   // Length based on data_ptr (Used for data_len)
      END_STRUCT;
      conf : Struct   // Configuration
         buffer_handler : Bool := TRUE;   // enable buffer handler
         halt : Bool;   // Halt exec. of queries.
      END_STRUCT;
      stat : Struct   // Status of last executed query
         done : Bool;   // Successfull
         error : Bool;   // Error, including timeout error
         busy : Bool;   // mb_master or mb_client is busy.
         error_comm : Bool;   // communication error (timeout or bad crc)
         status : Word;   // status word of mb_master or mb_client
      END_STRUCT;
      z : Struct   // Internal states
         q : Struct   // Query params
            mb_addr : UInt := 1;   // Station address
            mode : USInt := 0;   // Function code
            data_addr : UDInt;   // Data address
            data_len : UInt := 0;   // Data length
         END_STRUCT;
         run : Struct   // Constantly changing variables
            qid : UInt := 1;   // query id
            qid_cnt : UInt;   // Query id cnt. increase for each query, reset in controller. One loop each scan
            state : USInt;
            write : Bool;   // A write query is inserted
            discrete : Bool;
         END_STRUCT;
         sb : Struct   // Station block functionality
            sid : UInt;   // Device ID
            sid_cnt : UInt;   // Device id cnt
            sid_retry : UInt := 1;   // Retry device id, qComError
            retry_finished : Bool;
            head_insert : Bool;   // Inc. at mb_query on insert
            head_recive : Bool;   // Inc. at mb_query on rec.
            reset : Bool;
            log_data_addr : UDInt;   // Tmp.var. for transf. value to mb_device_footer
         END_STRUCT;
         buffer : Array[0..249] of Byte;
      END_STRUCT;
   END_VAR
   VAR_TEMP
      tLen : UInt;
      tPos : DInt;
      tDiscrete : Bool;
      "e" : Int;
      tBuffer : Array[0..249] of Byte;
   END_VAR
   VAR CONSTANT
      ORIGIN : USInt := 0;
      INSERT_QUERY : USInt := 1;
      INIT_QUERY : USInt := 2;
      EXEC_QUERY : USInt := 3;
      RECIVE_RESUALT : USInt := 4;
   END_VAR
BEGIN
   // Rexhip - Extended modbus library 
   // --- --- --- ---
   // License:  MIT-license
   // Author:   Ola Bjørnli
   // Web:      www.rexhip.com
   //           github.com/rexhip/rexhip
   // --- --- --- ---
   // 
   // For autmatic calculation of data_len, mb_query can only count whole
   // words (16 bits). This implices that the automatic length works well
   // for holding- and input registers, but dosen't work for dicreate
   // queries. For this queries data_len need to be specified manually.
   // After a query where data_len is specified, it need to be set back
   // to automatic. (#mb_query.data_len := #mb_query.c.auto_len;)
   //
   // Please read to the documentation and see the examples, before dive
   // into the code bellow.

   REGION Header            
       #Done := #Error := false;

       // qid_cnt is increased for every query (above) and reset back
       // to zero in mb_internal_e. Qid (query id) is increased when a
       // query finnish. A query will execute when qit_cnt = qid. Qid
       // is set back to "1" when all queryies has been executed.
       #z.run.qid_cnt += 1;
       IF #z.run.qid_cnt <> #z.run.qid
           OR #stat.busy // mb_master.busy or mb_client.busy
       THEN
           RETURN;
       END_IF;
   END_REGION

   REGION Pre-calc
       // Is this a discrete query ?
       CASE #mode OF
           1, 2, 5, 15: // Function codes
               #tDiscrete := true;
           200..202:
               CASE #data_addr OF
                   1..19999: // 1..9999, 10001..19999:
                       #tDiscrete := true;
               END_CASE;
       END_CASE;

       // data_len=0 => Automatically calculate the length.
       IF #data_len = 0 THEN
           #"e" := Serialize(SRC_VARIABLE := #data_ptr,
                           DEST_ARRAY => #tBuffer,
                           POS := #tPos);
           #tLen := DINT_TO_UINT
           (SEL(G := #tDiscrete, IN0 := #tPos / 2, IN1 := #tPos * 8));
       ELSE
           #tLen := #data_len;
       END_IF;
   END_REGION

   // Wait inserting next query if halted, else just continue.
   IF #z.run.state = #ORIGIN AND NOT #conf.halt THEN
       #z.run.state := #INSERT_QUERY;
   END_IF;

   CASE #z.run.state OF
       #INSERT_QUERY: // Transfer query params. to internal variables.

           // Figur out if this is a query that will write to the device.
           CASE #mode OF
               5, 6, 15, 16, 201, 202: // Write fc's.
                   #z.run.write := true;
               ELSE // Read
                   #z.run.write := false;
           END_CASE;

           #z.run.discrete := #tDiscrete;

           // The params is transfered over to the internal mem. They
           // are later transfered to the modbus master block or the
           // client block.
           #z.q.mb_addr := #mb_addr;
           #z.q.mode := #mode;
           #z.q.data_addr := #data_addr;
           #z.q.data_len := #tLen;

           IF #conf.buffer_handler AND #z.run.write THEN
               // Copy the content of #data_ptr to the buffer.
               #tPos := 0; // Start at the beginning of the buffer.
               #"e" := Serialize(SRC_VARIABLE := #data_ptr,
                               DEST_ARRAY => #z.buffer,
                               POS := #tPos);
           END_IF;
           // A msg. to station block foother FC, a new query has
           // been inserted.
           #z.sb.head_insert := true;

           #z.run.state := #INIT_QUERY; // State inside ctrl block.


       #RECIVE_RESUALT: // Query is finnished. (with or without error)  

           // Make sure that the query resault really belong to this
           // query. This may not be the case if another query before
           // is surrounded by a if-statement.
           IF #z.q.mb_addr = #mb_addr
               AND #z.q.mode = #mode
               AND #z.q.data_addr = #data_addr
               AND #z.q.data_len = #tLen
           THEN
               IF #stat.done // Successfull query (no error)
                   AND NOT #z.run.write  // If it's a read query.
                   AND #conf.buffer_handler
               THEN
                   // Copy the content from the buffer to #data_ptr
                   #tPos := 0; // Start at the beginning of the buffer.
                   #"e" := Deserialize(SRC_ARRAY := #z.buffer,
                                     DEST_VARIABLE => #data_ptr,
                                     POS := #tPos);
               END_IF;
               #Done := #stat.done;
               #Error := #stat.error;

               // Temperary store value, so it can be picked up
               // in the sb footer.
               #z.sb.log_data_addr := #data_addr;
               // Msg. to mb_station_footer.
               #z.sb.head_recive := true;
           END_IF;
           #z.run.qid += 1; // Next query
           #z.run.state := #ORIGIN; // (State before insert, see above)
   END_CASE;
END_FUNCTION_BLOCK

// folder: Library/Modbus/Core/Ctrl

FUNCTION_BLOCK "mb_master_1200_ctrl"   // FB90, SCL
{ S7_Optimized_Access := 'TRUE' }
VERSION : 1.0
   VAR_INPUT
      hardware_id : Port := 0;   // Hardware id
      baud : UDInt := 19200;   // Bits per second
   END_VAR
   VAR_OUTPUT
      Error : Bool;   // One or more errors in the whole application.
   END_VAR
   VAR_IN_OUT
      mb_query : "mb_query";
   END_VAR
   VAR
      conf : Struct   // Configuration that normal shouldn't need to be changed.
         parity : UInt := 2;   // 0=no-parity, 1=odd, 2=even.
         retries : USInt := 0;
         timeout_gain : Real := 2.0;   // Multiplied with the calculated value.
         timeout_offset : Time := T#0ms;   // Added to the calculated value.
      END_STRUCT;
      comm_load : MB_COMM_LOAD;
      master : MB_MASTER;
      buffer : "mb_internal_b";
      end : "mb_internal_e";   // FB common for both rtu and tcp.
   END_VAR
   VAR_TEMP
      tmp_err : Bool;
   END_VAR
   VAR CONSTANT
      INIT_QUERY : USInt := 2;
      EXEC_QUERY : USInt := 3;
      RECIVE_RESUALT : USInt := 4;
   END_VAR
BEGIN
   // Rexhip - Extended modbus library.
   // Please see top section of mb_query for more info.
   // 
   // RTU master for S7-1200
   // 
   // This FB use less memory then mb_master_1500_ctrl, but it only works for
   // S7-1200 PLC's. Please read the documentation, before dive into the code
   // bellow